screen "MTA-ALTAMC005" 1280x800, template "Plantilla-Alta-Cmp"
   Button "Botón_1" at 186,441 size 48x38; TextOff 'Incrementar'; Authorization "Operación"; PictureOff "Gráfico_3"
      on Press: SetBit("IncP5")
      on Release: ResetBit("IncP5")
   Button "Botón_2" at 186,401 size 48x38; TextOff 'Decrementar'; Authorization "Operación"; PictureOff "Gráfico_1"
      on Press: SetBit("DecP5")
      on Release: ResetBit("DecP5")
   Button "Botón_7" at 390,106 size 40x38; TextOff 'Text'; PictureOff "x"
      on Click: function_efd93a16()
   Button "Botón_8" at 310,600 size 96x35; TextOff 'Hecho'; Authorization "Administración de usuarios"
      on Press: SetTag("Varios_UltimoMantMC005_1", "HORAS5")
   TextField "Campo de texto_6" at 266,362 size 72x27; Text 'Seteada'
   TextField "Campo de texto_7" at 82,426 size 84x27; Text 'Prioridad'
   TextField "Campo de texto_8" at 362,363 size 40x27; Text 'Real'
   TextField "Campo de texto_11" at 26,343 size 158x27; Text 'Seteo de Prioridad'
   GraphicIOField "Campo ES gráfico_3" at 294,402 size 16x78; PictureList "BarraPrioridades"
      ProcessValue <- "VCMP5"
   GraphicIOField "Campo ES gráfico_5" at 374,402 size 16x78; PictureList "BarraPrioridades_1"
      ProcessValue <- "PriRealCMP5"
   SymbolicIOField "Campo ES simbólico_2" at 9,290 size 424x37; TextOff '0'; TextOn '1'; TextList "EstadoCmpAlta"
      ProcessValue <- "Est5"
      Visibility <- "MantMC005"
   TextField "Campo de texto_16" at 521,10 size 279x27; Text 'Menú Compresor ABC-5 (MC005)'
   TextField "Campo de texto_1" at 36,510 size 326x27; Text 'Tiempo de funcionamiento acumulado'
   TextField "Campo de texto_4" at 36,570 size 231x27; Text 'Próximo mantenimiento #1'
   TextField "Campo de texto_5" at 36,635 size 231x27; Text 'Próximo mantenimiento #2'
   Button "Botón_3" at 310,665 size 96x35; TextOff 'Hecho'; Authorization "Administración de usuarios"
      on Press: SetTag("Varios_UltimoMantMC005_2", "HORAS5")
   IOField "Campo ES_4" at 574,609 size 96x32; FormatPattern 99; Unit  min
      ProcessValue <- "DB-PurgaComAlta_Toff_PurgaABC5"
   IOField "Campo ES_5" at 574,654 size 96x32; FormatPattern 99; Unit  seg
      ProcessValue <- "DB-PurgaComAlta_Ton_PurgaABC5"
   TextField "Campo de texto_2" at 459,613 size 97x27; Text 'Tiempo Off'
   TextField "Campo de texto_3" at 459,655 size 96x27; Text 'Tiempo On'
   Switch "Interruptor_2" at 459,548 size 120x40; TextOff 'OFF'; CaptionText 'Switch'; TextOn 'ON'
      ProcessValue <- "DB-PurgaComAlta_Habil_PurgaABC5"
   Button "Botón_4" at 595,548 size 80x40; TextOff 'Prueba'
      on Press: SetBit("DB-PurgaComAlta_Prueba_PurgaABC5")
      on Release: ResetBit("DB-PurgaComAlta_Prueba_PurgaABC5")
      Appearance <- "MC005_EVP"
      ObjectEnable <- "MC005_EVP"
   TextField "Campo de texto_9" at 456,510 size 131x27; Text 'Ciclo de Purga:'
   GraphicIOField "Campo ES gráfico_2" at 10,280 size 422x6; PictureList "Indicador"
      ProcessValue <- "AnimMotorMC005"
   SymbolicIOField "Campo ES simbólico_4" at 19,246 size 290x21; TextOff '0'; TextOn '1'; TextList "EstadoMotor"
      ProcessValue <- "AnimMotorMC005"
   Button "Botón_6" at 13,154 size 88x62; TextOff 'ABC 5'
   Switch "Interruptor_1" at 150,167 size 37x37; TextOn '1'; TextOff '0'; CaptionText 'Switch'; PictureOff "A2"; Authorization "Operación"; PictureOn "A"
      ProcessValue <- "Auto5"
      Visibility <- "MantMC005"
   ScreenModuleView "Faceplate_6_1" at 342,236 size 76x34; ScreenModuleType ""
      Guid_{11997190-52606} <- "IndV5"
      Guid_{11997190-52610} <- "IndR5"
      Guid_{11997190-52608} <- "IndVparp5"
   ScreenModuleView "Faceplate_7_1" at 213,158 size 207x70
      Guid_{11997190-23983} <- "ParadaMC005"
      Guid_{11997190-23981} <- "MarchaMC005"
      Guid_{11997190-90329} <- "ForzarParada5"
      Guid_{11997190-180841} <- "MantMC005"
      Guid_{11997190-89807} <- "SPOFFF5"
      Guid_{11997190-89795} <- "ForzandoMarcha5"
      Guid_{11997190-90325} <- "MarchaMC005"
      Guid_{11997190-88662} <- "MarchaOK5"
      Guid_{11997190-23985} <- "AnimMenuMC005"
      Guid_{11997190-89805} <- "SPONF5"
   IOField "Campo ES_7" at 24,535 size 173x35; Authorization "Administración de usuarios"; FormatPattern 999999999; Unit  hs
      ProcessValue <- "HORAS5"
      Appearance <- "EstadoMantMC005"
   IOField "Campo ES_1" at 204,535 size 80x35; Authorization "Administración de usuarios"; FormatPattern 99; Unit  min
      ProcessValue <- "MIN5"
   IOField "Campo ES_2" at 24,595 size 173x35; FormatPattern 999999999; Unit  hs
      ProcessValue <- "ProxMantMC005_1"
      Appearance <- "LimiteMantMC005_1"
   IOField "Campo ES_3" at 24,660 size 173x35; FormatPattern 999999999; Unit  hs
      ProcessValue <- "ProxMantMC005_2"
      Appearance <- "LimiteMantMC005_2"

screen "MTA-Avisos" 1280x800, template "Plantilla"
   AlarmView "Visor de avisos_1" at 61,61 size 1174x631
   TextField "Campo de texto_16" at 613,9 size 54x27; Text 'Avisos'

screen "MTA-Avisos-Histórico" 1280x800, template "Plantilla"
   AlarmView "Visor de avisos_1" at 61,61 size 1174x631; AlarmLog "Fichero de avisos_MTA"
   TextField "Campo de texto_16" at 573,9 size 157x27; Text 'Histótico de Avisos'

screen "MTA-AyudaCFG1" 1280x800, template "Plantilla"
   TextField "Campo de texto_1" at 66,128 size 540x220; Text 'Cada compresor tiene su banda de presiones. Las 5 bandas para los 5 compresores se encuentran desfasadas una cantidad, determinada por el parámetro “Separación de presión entre bandas de presión de regulación”. Las posiciones de las bandas están determinadas por las prioridades. La banda de más arriba es la de Prioridad 1, y la de más abajo es la de prioridad 5. Los cambios en las prioridades que se le asignan a cada compresor no alteran el orden de las bandas de regulación. Las bandas siempre tienen el orden en función de las prioridades: la banda de más arriba es la de Prioridad 1, le sigue la 2, la 3 , la 4 y la de más abajo es la de prioridad 5.'
   TextField "Campo de texto_2" at 42,112 size 507x27; Text 'Posición de las bandas de regulación y parámetros a ajustar'
   TextField "Campo de texto_3" at 66,416 size 508x220; Text 'Cuando la presión medida se encuentre por deajo de la presión crítica inferior, cualquier compresor que se ponga en marcha comenzará a funcionar independientemente de si existen o no sopladoras encendidas. Una vez que la presión haya regresado a su nivel normal (es decir, que haya superado el valor de “Presión Crítica Superior”), los compresores regularán de manera normal, y se encenderán únicamente si existen sopladoras encendidas. La utilidad de este comportamiento, es que permite recuperar rápidamente la presión en casos tales como cuando por largo tiempo los compresores y sopladoras estuvieron apagados, y las pérdidas en las cañerías hicieron que la presión llegara a cero o a un valor cercano'
   TextField "Campo de texto_4" at 42,400 size 235x27; Text 'Utilidad de la presión crítica'
   TextField "Campo de texto_5" at 905,92 size 123x32; Text 'Banda de regulación Compresor Prioridad 1'
   TextField "Campo de texto_6" at 905,172 size 123x32; Text 'Banda de regulación Compresor Prioridad 2'
   TextField "Campo de texto_7" at 905,252 size 123x32; Text 'Banda de regulación Compresor Prioridad 3'
   TextField "Campo de texto_8" at 905,332 size 123x32; Text 'Banda de regulación Compresor Prioridad 4'
   TextField "Campo de texto_9" at 905,412 size 123x32; Text 'Banda de regulación Compresor Prioridad 5'
   TextField "Campo de texto_11" at 1148,498 size 88x32; Text 'Presión mínima para regulación'
   TextField "Campo de texto_12" at 708,557 size 128x18; Text 'Presión Crítica Superior'
   TextField "Campo de texto_13" at 708,611 size 122x18; Text 'Presión Crítica Inferior'
   TextField "Campo de texto_14" at 1162,199 size 85x46; Text 'Histéresis para regulación de presión'
   TextField "Campo de texto_15" at 658,199 size 140x46; Text 'Separación de presiones entre bandas de regulación de presión'
   Button "Botón_12" at 1089,638 size 160x49; TextOff 'Volver'
      on Click: ActivateScreen("MTA-CFGALTA", 0)
   TextField "Campo de texto_16" at 414,9 size 455x27; Text 'Ayuda: Configuración modo AUTO (Compresores Alta)'
   TextField "Campo de texto_10" at 905,492 size 123x32; Text 'Banda de regulación Compresor Prioridad 5'

screen "MTA-AyudaCmpAlta" 1280x800, template "Plantilla"
   Switch "Interruptor_1" at 1192,363 size 40x40; TextOn '1'; TextOff '0'; CaptionText 'Switch'; PictureOff "MECH2"; PictureOn "MECH1"
      ProcessValue <- "CERO"
   GraphicIOField "Campo ES gráfico_6" at 763,381 size 9x45; PictureList "BarraPrioridades"
      ProcessValue <- "VCMP3"
      Visibility <- "MantMC003"
   GraphicIOField "Campo ES gráfico_9" at 772,381 size 9x45; PictureList "BarraPrioridades_1"
      ProcessValue <- "PriRealCMP3"
      Visibility <- "MantMC003"
   GraphicView "Visor de gráficos_1" at 660,384 size 28x27; Picture "A2"
   TextField "Campo de texto_6" at 285,315 size 125x61; Text 'Estado del motor del Compresor'
   TextField "Campo de texto_10" at 413,297 size 113x61; Text 'Nombre del Compresor'
   TextField "Campo de texto_1" at 532,218 size 108x80; Text 'Estado lógico del Compresor (Programa)'
   GraphicView "Visor de gráficos_3" at 694,382 size 28x30; Picture "PilotLight_Round_GN_On_256c"
   GraphicView "Visor de gráficos_4" at 726,382 size 28x30; Picture "PilotLight_Round_RN_Off_256c"
   GraphicView "Visor de gráficos_5" at 126,91 size 28x30; Picture "PilotLight_Round_GN_Off_256c"
   GraphicView "Visor de gráficos_7" at 94,91 size 28x30; Picture "PilotLight_Round_RN_Off_256c"
   GraphicView "Visor de gráficos_8" at 126,131 size 28x30; Picture "PilotLight_Round_GN_Off_256c"
   GraphicView "Visor de gráficos_9" at 94,131 size 28x30; Picture "PilotLight_Round_RN_On_256c"
   GraphicView "Visor de gráficos_10" at 126,171 size 28x30; Picture "PilotLight_Round_GN_Off_256c"
   GraphicView "Visor de gráficos_11" at 94,171 size 28x30; Picture "PilotLight_Round_RN_On_256c"
   GraphicView "Visor de gráficos_12" at 126,211 size 28x30; Picture "PilotLight_Round_GN_On_256c"
   GraphicView "Visor de gráficos_13" at 94,211 size 28x30; Picture "PilotLight_Round_RN_Off_256c"
   GraphicView "Visor de gráficos_14" at 126,171 size 28x30; Picture "PilotLight_Round_GN_On_256c"
   GraphicIOField "Plantilla_Campo ES gráfico_5" at 897,433 size 65x60; PictureList "Motor2"
      ProcessValue <- "UNO"
   GraphicView "Visor de gráficos_2" at 924,363 size 260x142; Picture "ALTA1_1"
   GraphicView "Visor de gráficos_6" at 971,83 size 262x142; Picture "LOCAl"
   TextField "Campo de texto_7" at 607,463 size 54x42; Text 'Manual'
   TextField "Campo de texto_11" at 1067,286 size 199x76; Text 'El modo local transfiere el control del Compresor a su panel original'
   TextField "Campo de texto_12" at 1056,264 size 210x42; Text 'Activación de modo "LOCAL"'
   TextField "Campo de texto_13" at 695,98 size 210x42; Text 'Indicación de modo "LOCAL"'
   TextField "Campo de texto_16" at 926,529 size 134x42; Text 'Código de Colores'
   TextField "Campo de texto_18" at 529,9 size 241x27; Text 'Ayuda: Compresores de Alta'
   TextField "Campo de texto_3" at 703,239 size 90x80; Text 'Prioridad de arranque Seteada'
   TextField "Campo de texto_4" at 815,215 size 95x80; Text 'Prioridad de arranque Actual'
   TextField "Campo de texto_5" at 700,485 size 129x61; Text 'Horas de marcha acumuladas'
   TextField "Campo de texto_2" at 223,92 size 170x42; Text 'Deshabilitado / En Falla'
   TextField "Campo de texto_8" at 223,132 size 284x42; Text 'Habilitado y Parado / Sin requerimiento'
   TextField "Campo de texto_9" at 223,172 size 268x42; Text 'Parado con Requerimiento de Marcha'
   TextField "Campo de texto_14" at 223,212 size 122x42; Text 'En Vacío / Carga'
   TextField "Campo de texto_15" at 561,383 size 61x22; Text 'En carga'
   Button "Botón_3" at 95,559 size 280x70; TextOff 'Ayuda de Manejo'; PictureOff "x"
      on Click: ActivateScreen("MTA-AyudaCmpAlta_1", 0)
   GraphicIOField "Campo ES gráfico_4" at 421,438 size 374x6; PictureList "Indicador"
      ProcessValue <- "UNO"
   SymbolicIOField "Campo ES simbólico_4" at 440,410 size 178x21; TextOff '0'; TextOn '1'; TextList "EstadoMotor"
      ProcessValue <- "UNO"
   TextField "Campo de texto_19" at 434,377 size 66x32; Text 'ABC 2'
   IOField "Campo ES_6" at 662,413 size 85x19; FormatPattern 999999999; Unit  hs

screen "MTA-AyudaCmpAlta_1" 1280x800, template "Plantilla"
   TextField "Campo de texto_18" at 529,9 size 241x27; Text 'Ayuda: Compresores de Alta'
   TextField "Campo de texto_5" at 466,549 size 701x99; Text 'Para poder resetear las horas acumuladas de cada compresor se requiere clave de administrador. Si la cantidad máxima de horas es superada se generará un aviso y el indicador de horas se pondrá de color rojo. Para eliminar este aviso se deben resetear la cantidad de horas acumuladas, y se debería considerar la posibilidad de bajar la prioridad del compresor.'
   TextField "Campo de texto_1" at 286,362 size 72x27; Text 'Seteada'
   TextField "Campo de texto_2" at 102,426 size 84x27; Text 'Prioridad'
   TextField "Campo de texto_10" at 382,363 size 40x27; Text 'Real'
   TextField "Campo de texto_6" at 46,520 size 326x27; Text 'Tiempo de funcionamiento acumulado'
   TextField "Campo de texto_3" at 46,343 size 158x27; Text 'Seteo de Prioridad'
   Button "Botón_1" at 206,442 size 48x38; TextOff 'Incrementar'; Authorization "Operación"; PictureOff "Gráfico_3"
   Button "Botón_2" at 206,402 size 48x38; TextOff 'Decrementar'; Authorization "Operación"; PictureOff "Gráfico_1"
   Button "Botón_3" at 410,106 size 40x38; TextOff 'Text'; PictureOff "x"
      on Click: function_efd93a16()
   Button "Botón_4" at 320,558 size 96x70; TextOff 'Reset'; Authorization "Administración de usuarios"
   GraphicIOField "Campo ES gráfico_1" at 314,402 size 16x78; PictureList "BarraPrioridades"
      ProcessValue <- "VCMP2"
   GraphicIOField "Campo ES gráfico_2" at 394,402 size 16x78; PictureList "BarraPrioridades_1"
      ProcessValue <- "PriRealCMP2"
   TextField "Campo de texto_4" at 466,381 size 709x80; Text 'Para poder cambiar las prioridades de un compresor se requiere que todas las soplatoras estén desactivadas. No habrá ningúna modificación en la cantidad de compresores requeridos si el ajuste de prioridades se realiza en un tiempo menor al "Tiempo de apagado de sopladoras". Una vez terminado el ajuste el usuario debería activar nuevamente las sopladoras correspondientes.'
   TextField "Campo de texto_7" at 466,150 size 658x61; Text 'Modo MANUAL: El motor del compresor se acciona con los pulsadores de marcha y parada. El rango de presiones en el cual el compresor estará en carga debe ser seteado (On: entra en carga / Off: sale de carga) y es independiente para cada compresor.'
   TextField "Campo de texto_8" at 466,222 size 812x99; Text 'Modo AUTO: El motor del compresor va a requerir marcha de acuerdo con la cantidad de compresores necesarios para las sopladoras que estén activas. El rango de presiones en el cual el compresor estará en carga depende de su prioridad real. El compresor puede entrar en carga / requerir marcha de manera extraordinaria si la presión de la linea es menor que la "Presión Crítica" estando en modo AUTOMÁTICO.'
   TextField "Campo de texto_9" at 202,296 size 76x27; Text 'En Vacío'
   GraphicIOField "Campo ES gráfico_3" at 30,279 size 422x6; PictureList "Indicador"
      ProcessValue <- "UNO"
   SymbolicIOField "Campo ES simbólico_2" at 39,245 size 290x21; TextOff '0'; TextOn '1'; TextList "EstadoMotor"
      ProcessValue <- "UNO"
   Button "Botón_6" at 41,153 size 88x62; TextOff 'ABC 3'
   Switch "Interruptor_1" at 170,166 size 37x37; TextOn '1'; TextOff '0'; CaptionText 'Switch'; PictureOff "A2"; PictureOn "A"
      ProcessValue <- "Auto1"
      Visibility <- "MantMC002"
   ScreenModuleView "Faceplate_7_1" at 241,157 size 200x70
      Guid_{11997190-23985} <- "AnimMenuMC001"
   IOField "Campo ES_7" at 88,558 size 173x35; FormatPattern 999999999; Unit  hs
   IOField "Campo ES_1" at 103,590 size 173x35; FormatPattern 999999999; Unit  min
   GraphicView "Visor de gráficos_12" at 356,232 size 36x38; Picture "PilotLight_Round_GN_On_256c"
   GraphicView "Visor de gráficos_13" at 396,232 size 36x38; Picture "PilotLight_Round_RN_Off_256c"

screen "MTA-AyudaColores" 1280x800, template "Plantilla"
   GraphicView "Visor de gráficos_1" at 156,507 size 64x58; Picture "indAmarillo"
   GraphicView "Visor de gráficos_3" at 156,251 size 64x58; Picture "indCeleste"
   GraphicView "Visor de gráficos_4" at 156,315 size 64x58; Picture "indDorado"
   GraphicView "Visor de gráficos_5" at 156,187 size 64x58; Picture "indGris"
   GraphicView "Visor de gráficos_6" at 156,379 size 64x58; Picture "indRojo"
   GraphicView "Visor de gráficos_7" at 156,443 size 64x58; Picture "indVerde"
   TextField "Campo de texto_1" at 234,518 size 172x42; Text 'Sobrecarga de corriente'
   TextField "Campo de texto_2" at 130,112 size 233x32; Text 'Codificación de colores'
   TextField "Campo de texto_3" at 234,262 size 75x42; Text 'Habilitado'
   TextField "Campo de texto_4" at 234,326 size 431x42; Text 'Detenido (en algunos casos también significa modo manual)'
   TextField "Campo de texto_5" at 234,198 size 99x42; Text 'Deshabilitado'
   TextField "Campo de texto_6" at 234,390 size 56x42; Text 'En falla'
   TextField "Campo de texto_7" at 234,454 size 77x42; Text 'En Marcha'
   TextField "Campo de texto_8" at 130,598 size 666x58; Text 'Los colores indican los estados de los motores / compresores / secadores de manera rápida. La codificación de colores siempre está acompañada de un texto que contiene la misma información.'
   TextField "Campo de texto_9" at 130,646 size 1002x40; Text 'En algunos casos también aparecen los colores Verde Oscuro y Azul Oscuro que indican los estados de "Arrancando" y "Deteniéndose" respectivamente.'
   TextField "Campo de texto_16" at 542,9 size 200x27; Text 'Ayuda: Estados/Colores'

screen "MTA-AyudaMotores" 1280x800, template "Plantilla"
   TextField "Campo de texto_5" at 159,478 size 343x42; Text 'Representación de Motor con código de colores'
   TextField "Campo de texto_8" at 50,294 size 461x58; Text 'La Deshabilitación del motor provoca también la detención del mismo. La Habilitación del motor permite operar el pulsador de Marcha.'
   TextField "Campo de texto_9" at 882,291 size 279x58; Text 'Para poder marchar el motor es necesario que el mismo esté habilitado'
   GraphicView "Visor de gráficos_2" at 624,407 size 64x103; Picture "Bomba"
   GraphicIOField "Plantilla_Campo ES gráfico_4" at 660,481 size 81x68; PictureList "Motor2"
      ProcessValue <- "UNO"
   SymbolicIOField "Campo ES simbólico_3" at 572,220 size 220x29; TextOff '0'; TextOn '1'; TextList "EstadoMotor"
      ProcessValue <- "UNO"
   TextField "Campo de texto_10" at 575,161 size 52x23; Text 'MP013'
   TextField "Campo de texto_17" at 573,193 size 146x18; Text 'Chillers Envasado - Backup'
   ScreenModuleView "ControlMotor-NoAUTO_4" at 599,262 size 171x108
   TextField "Campo de texto_1" at 39,261 size 436x42; Text 'Habilitación/Deshabilitación del accionamiento desde el panel'
   TextField "Campo de texto_2" at 871,261 size 179x42; Text 'Orden de Marchar motor'
   TextField "Campo de texto_3" at 871,373 size 160x42; Text 'Orden de Parar motor'
   TextField "Campo de texto_4" at 119,205 size 376x42; Text 'Estado del motor (descripción del código de colores)'
   TextField "Campo de texto_6" at 871,165 size 251x23; Text 'Nombre simbólico en el programa'
   TextField "Campo de texto_7" at 871,197 size 135x42; Text 'Nombre del motor'
   TextField "Campo de texto_16" at 573,9 size 135x27; Text 'Ayuda: Motores'

screen "MTA-AyudaSecAlta" 1280x800, template "Plantilla"
   GraphicIOField "Campo ES gráfico_1" at 141,455 size 511x6; PictureList "Indicador"
      ProcessValue <- "UNO"
   GraphicIOField "Campo ES gráfico_2" at 141,639 size 511x6; PictureList "Indicador"
      ProcessValue <- "CERO"
   GraphicIOField "Campo ES gráfico_7" at 962,373 size 309x81; PictureList "Secador2"
      ProcessValue <- "UNO"
   GraphicView "Visor de gráficos_2" at 988,283 size 260x142; Picture "secador3_1"
   GraphicView "Visor de gráficos_6" at 971,83 size 262x142; Picture "secador3d_1"
   GraphicView "Visor de gráficos_1" at 318,376 size 35x35; Picture "A2"
   GraphicView "Visor de gráficos_3" at 318,562 size 35x35; Picture "A"
   GraphicView "Visor de gráficos_5" at 414,369 size 202x78; Picture "menu2"
   GraphicView "Visor de gráficos_7" at 413,552 size 231x79; Picture "menu3"
   TextField "Campo de texto_8" at 290,158 size 333x94; Text 'La Deshabilitación del Secador provoca también la detención del mismo. La Habilitación del Secador permite su operaración desde el panel.'
   TextField "Campo de texto_9" at 474,275 size 211x76; Text 'Para poder marchar el Secador es necesario que el mismo esté habilitado'
   TextField "Campo de texto_3" at 279,133 size 203x42; Text 'Habilitación/Deshabilitación'
   TextField "Campo de texto_4" at 463,245 size 192x42; Text 'Orden de Marchar Secador'
   TextField "Campo de texto_5" at 679,495 size 173x42; Text 'Orden de Parar Secador'
   TextField "Campo de texto_6" at 53,267 size 143x42; Text 'Estado del Secador'
   TextField "Campo de texto_7" at 303,295 size 54x42; Text 'Manual'
   TextField "Campo de texto_10" at 175,309 size 91x61; Text 'Nombre del Secador'
   TextField "Campo de texto_11" at 706,275 size 180x76; Text 'El modo local transfiere el control del Secador a su panel original'
   TextField "Campo de texto_12" at 695,245 size 210x42; Text 'Activación de modo "LOCAL"'
   TextField "Campo de texto_13" at 695,98 size 210x42; Text 'Indicación de modo "LOCAL"'
   TextField "Campo de texto_14" at 714,643 size 520x76; Text 'Cada Secador puede relacionar su estado con uno o dos compresores de alta. Mientras alguno de los compresores seleccionados esté en marcha, el secador se mantendrá en funcionamiento.'
   TextField "Campo de texto_15" at 703,613 size 255x42; Text 'Enclavamientos (Modo Automático)'
   TextField "Campo de texto_16" at 1062,513 size 134x42; Text 'Código de Colores'
   TextField "Campo de texto_17" at 310,487 size 38x42; Text 'Auto'
   TextField "Campo de texto_18" at 529,9 size 219x27; Text 'Ayuda: Secadores de Alta'
   TextField "Campo de texto_1" at 166,377 size 89x39; Text 'ABC 2'
   SymbolicIOField "Campo ES simbólico_1" at 168,413 size 242x21; TextOff '0'; TextOn '1'; TextList "EstadoMotor"
      ProcessValue <- "UNO"
   TextField "Campo de texto_2" at 166,561 size 89x39; Text 'ABC 2'
   SymbolicIOField "Campo ES simbólico_2" at 168,597 size 242x21; TextOff '0'; TextOn '1'; TextList "EstadoMotor"
      ProcessValue <- "CERO"
   Switch "Interruptor_1" at 928,331 size 40x40; TextOn '1'; TextOff '0'; CaptionText 'Switch'; PictureOff "MECH2"; PictureOn "MECH1"
      ProcessValue <- "CERO"

screen "MTA-AyudaSecBaja" 1280x800, template "Plantilla"
   GraphicIOField "Campo ES gráfico_3" at 626,509 size 510x6; PictureList "Indicador"
      ProcessValue <- "UNO"
   GraphicIOField "Campo ES gráfico_8" at 303,471 size 269x90; PictureList "BaseSullChico"
      ProcessValue <- "UNO"
   GraphicView "Visor de gráficos_1" at 336,357 size 201x179; Picture "secador_1"
   GraphicView "Visor de gráficos_3" at 344,125 size 201x179; Picture "Copia de secador"
   TextField "Campo de texto_11" at 50,363 size 180x76; Text 'El modo local transfiere el control del Secador a su panel original'
   TextField "Campo de texto_12" at 39,333 size 210x42; Text 'Activación de modo "LOCAL"'
   GraphicView "Visor de gráficos_5" at 917,426 size 202x78; Picture "menu2"
   TextField "Campo de texto_2" at 95,141 size 210x42; Text 'Indicación de modo "LOCAL"'
   TextField "Campo de texto_5" at 643,433 size 107x39; Text 'Sullair 1'
   TextField "Campo de texto_7" at 650,472 size 54x23; Text 'Marcha'
   TextField "Campo de texto_8" at 802,214 size 333x94; Text 'La Deshabilitación del Secador provoca también la detención del mismo. La Habilitación del Secador permite su operaración desde el panel.'
   TextField "Campo de texto_9" at 986,331 size 211x76; Text 'Para poder marchar el Secador es necesario que el mismo esté habilitado'
   TextField "Campo de texto_4" at 791,189 size 203x42; Text 'Habilitación/Deshabilitación'
   TextField "Campo de texto_10" at 975,301 size 192x42; Text 'Orden de Marchar Secador'
   TextField "Campo de texto_13" at 1031,559 size 173x42; Text 'Orden de Parar Secador'
   TextField "Campo de texto_14" at 564,558 size 143x42; Text 'Estado del Secador'
   TextField "Campo de texto_15" at 655,365 size 91x61; Text 'Nombre del Secador'
   TextField "Campo de texto_16" at 529,9 size 224x27; Text 'Ayuda: Secadores de Baja'
   Switch "Interruptor_8" at 275,422 size 40x40; TextOn '1'; TextOff '0'; CaptionText 'Switch'; PictureOff "MECH2"; PictureOn "MECH1"

screen "MTA-AyudaVentiladores" 1280x800, template "Plantilla"
   GraphicIOField "Campo ES gráfico_6" at 328,342 size 511x6; PictureList "Indicador"
      ProcessValue <- "CERO"
   TextField "Campo de texto_5" at 957,566 size 184x61; Text 'Representación de Motor con código de colores'
   TextField "Campo de texto_8" at 218,134 size 461x58; Text 'La Deshabilitación del motor provoca también la detención del mismo. La Habilitación del motor permite operarlo desde el panel.'
   TextField "Campo de texto_9" at 818,131 size 279x58; Text 'Para poder marchar el motor es necesario que el mismo esté habilitado'
   TextField "Campo de texto_1" at 207,101 size 436x42; Text 'Habilitación/Deshabilitación del accionamiento desde el panel'
   TextField "Campo de texto_2" at 807,101 size 179x42; Text 'Orden de Marchar motor'
   TextField "Campo de texto_4" at 197,542 size 250x61; Text 'Estado del motor (descripción del código de colores)'
   TextField "Campo de texto_7" at 107,251 size 135x42; Text 'Nombre del motor'
   GraphicView "Visor de gráficos_3" at 508,439 size 242x85; Picture "menu4_1"
   GraphicView "Visor de gráficos_4" at 508,253 size 226x85; Picture "menu2"
   GraphicView "Visor de gráficos_5" at 473,452 size 29x29; Picture "A"
   GraphicView "Visor de gráficos_6" at 473,268 size 29x29; Picture "A2"
   TextField "Campo de texto_12" at 957,478 size 156x61; Text 'Indicación ventilador en Marcha'
   TextField "Campo de texto_13" at 957,310 size 156x61; Text 'Indicación ventilador Detenido'
   TextField "Campo de texto_3" at 793,372 size 160x42; Text 'Orden de Parar motor'
   TextField "Campo de texto_6" at 413,638 size 729x61; Text 'Modo Automático Cada ventilador se pondrá en Marcha si la temperatura del agua sensada se encuentra por encima del valor de "On" y se apagará una vez que esté por debajo del valor de "Off"'
   TextField "Campo de texto_14" at 464,385 size 38x23; Text 'Auto'
   TextField "Campo de texto_15" at 448,209 size 54x23; Text 'Manual'
   TextField "Campo de texto_16" at 556,9 size 171x27; Text 'Ayuda: Ventiladores'
   TextField "Campo de texto_11" at 337,268 size 126x32; Text 'Ventilador 3'
   SymbolicIOField "Campo ES simbólico_1" at 339,304 size 170x21; TextOff '0'; TextOn '1'; TextList "EstadoMotor"
      ProcessValue <- "CERO"
   GraphicIOField "Campo ES gráfico_1" at 328,524 size 511x6; PictureList "Indicador"
      ProcessValue <- "UNO"
   TextField "Campo de texto_10" at 337,452 size 126x32; Text 'Ventilador 3'
   SymbolicIOField "Campo ES simbólico_2" at 339,488 size 170x21; TextOff '0'; TextOn '1'; TextList "EstadoMotor"
      ProcessValue <- "UNO"
   GraphicView "Visor de gráficos_18" at 757,262 size 71x70; Picture "Vent1"
   GraphicView "Visor de gráficos_1" at 757,446 size 71x70; Picture "Vent1"
   GraphicView "Visor de gráficos_2" at 757,446 size 71x70; Picture "Vent2"

screen "MTA-Booster" 1280x800, template "Plantilla"
   IOField "Campo ES_19" at 28,357 size 90x23; FormatPattern 999999999; Unit  hs
      ProcessValue <- "ProxMantBoost1"
      Appearance <- "LimiteMantBoost1"
   IOField "Campo ES_17" at 1109,356 size 90x23; FormatPattern 999999999; Unit  hs
      ProcessValue <- "ProxMantBoost2"
      Appearance <- "LimiteMantBoost2"
   GraphicView "Visor de gráficos_3" at 185,341 size 300x202; Picture "Booster-A"
   TextField "Campo de texto_16" at 0,10 size 1280x27; Text 'Boosters'
   GraphicIOField "Campo ES gráfico_1" at 238,431 size 64x70; PictureList "Motor Grande"
      ProcessValue <- "AnimaMotBooster"
   GraphicIOField "Campo ES gráfico_2" at 364,296 size 34x52; PictureList "Motor Chico"
      ProcessValue <- "AnimaMotBooster"
   GraphicIOField "Campo ES gráfico_3" at 208,410 size 221x101; PictureList "Hélice"
      ProcessValue <- "Booster_Conf_Marcha"
   SymbolicIOField "Campo ES simbólico_1" at 949,53 size 322x37; TextOff '0'; TextOn '1'; TextList "Presostato Ctrl"
      Appearance <- "Booster_Presost_Ctrl"
      ProcessValue <- "Booster_Presost_Ctrl"
   SymbolicIOField "Campo ES simbólico_2" at 949,95 size 321x37; TextOff '0'; TextOn '1'; TextList "Presostato de Alarma"
      ProcessValue <- "Booster_Presost_PA"
      Appearance <- "Booster_Presost_PA"
   GraphicView "Visor de gráficos_4" at 761,341 size 300x202; Picture "Booster-A"
   GraphicIOField "Campo ES gráfico_4" at 814,431 size 64x70; PictureList "Motor Grande"
      ProcessValue <- "AnimaMotBooster2"
   GraphicIOField "Campo ES gráfico_5" at 940,296 size 34x52; PictureList "Motor Chico"
      ProcessValue <- "AnimaMotBooster2"
   GraphicIOField "Campo ES gráfico_6" at 784,410 size 221x101; PictureList "Hélice"
      ProcessValue <- "Booster2_Conf_Marcha"
   GraphicView "Visor de gráficos_2" at 460,408 size 40x40; Picture "MECH2"
   GraphicView "Visor de gráficos_1" at 460,408 size 40x40; Picture "MECH1"
      Visibility <- "Booster_ModoManten"
   Button "Botón_6" at 460,408 size 40x40; TextOff 'Text'; PictureList "Mantenimiento"
      on Release: SetBit("Booster_PlsManten")
   IOField "Campo ES_1" at 217,338 size 90x23; Authorization "Administración de usuarios"; FormatPattern 999999999; Unit  hs.
      ProcessValue <- "HorasBoost1"
      Appearance <- "LimiteMantBoost1"
   IOField "Campo ES_2" at 790,338 size 90x23; Authorization "Administración de usuarios"; FormatPattern 999999999; Unit  hs.
      ProcessValue <- "HorasBoost2"
      Appearance <- "LimiteMantBoost2"
   Switch "Interruptor_2" at 361,96 size 72x40; TextOff 'No'; CaptionText 'Switch'; TextOn 'Si'
      ProcessValue <- "BoostPrHoras"
   TextField "Campo de texto_1" at 25,103 size 312x23; Text 'Control de Prioridades por horas de Marcha'
   Button "Botón_1" at 518,484 size 185x39; TextOff 'Invertir Prioridades'
      on Click: SetBit("BoostInvPMan")
      Visibility <- "BoostPrHoras"
   IOField "Campo ES_3" at 359,151 size 130x31; FormatPattern 99999; Unit  hs.
      ProcessValue <- "DifHorINVBoost"
      Visibility <- "BoostPrHoras"
   TextField "Campo de texto_2" at 241,152 size 93x23; Text 'Invertir cada'
      Visibility <- "BoostPrHoras"
   IOField "Campo ES_4" at 359,191 size 130x31; FormatPattern 99999; Unit  min.
      ProcessValue <- "TiempoAyudaON"
   TextField "Campo de texto_3" at 78,192 size 255x23; Text 'Tiempo para ayuda Booster auxiliar'
   IOField "Campo ES_5" at 359,231 size 130x31; FormatPattern 99999; Unit  seg.
      ProcessValue <- "TiempoAyudaOFF"
   TextField "Campo de texto_4" at 61,232 size 273x23; Text 'Tiempo para apagado Booster auxiliar'
   TextField "Campo de texto_5" at 187,550 size 250x27; Text 'Prioridad Marcha 2'
   TextField "Campo de texto_6" at 762,550 size 250x27; Text 'Prioridad Marcha 2'
   Button "Botón_7" at 849,639 size 100x27; TextOff 'Manual'
      on Release: SetBit("Booster2_PlsManual")
      Appearance <- "Booster2_ModoManual"
   Button "Botón_8" at 849,607 size 100x27; TextOff 'Automático'
      on Release: SetBit("Booster2_PlsAutoma")
      Appearance <- "Booster2_ModoAutoma"
   Button "Botón_9" at 960,607 size 96x27; TextOff 'Encender'; TextOn 'Encendido'
      on Release: SetBit("Booster2OrdMarcha")
      Appearance <- "Booster2_Conf_Marcha"
   Button "Botón_10" at 960,639 size 96x27; TextOff 'Detener'
      on Release: ResetBit("Booster2OrdMarcha")
   Switch "Interruptor_3" at 730,607 size 96x59; TextOff 'Deshabilitado'; CaptionText 'Habilitacion'; TextOn 'Habilitado'
      ProcessValue <- "Booster2_Habilitacion"
   GraphicView "Visor de gráficos_5" at 1036,408 size 40x40; Picture "MECH2"
   GraphicView "Visor de gráficos_6" at 1036,408 size 40x40; Picture "MECH1"
      Visibility <- "Booster2_ModoManten"
   Button "Botón_11" at 1036,408 size 40x40; TextOff 'Text'; PictureList "Mantenimiento"
      on Release: SetBit("Booster2_PlsManten")
   Button "Botón_2" at 275,639 size 96x27; TextOff 'Manual'
      on Release: SetBit("Booster_PlsManual")
      Appearance <- "Booster_ModoManual"
   Button "Botón_3" at 275,607 size 96x27; TextOff 'Automático'
      on Release: SetBit("Booster_PlsAutoma")
      Appearance <- "Booster_ModoAutoma"
   Button "Botón_5" at 384,607 size 96x27; TextOff 'Encender'; TextOn 'Encendido'
      on Release: SetBit("BoosterOrdMarcha")
      Appearance <- "Booster_Conf_Marcha"
   Button "Botón_4" at 384,639 size 96x27; TextOff 'Detener'
      on Release: ResetBit("BoosterOrdMarcha")
   Switch "Interruptor_1" at 153,607 size 96x59; TextOff 'Deshabilitado'; CaptionText 'Habilitacion'; TextOn 'Habilitado'
      ProcessValue <- "Booster_Habilitacion"
   IOField "Campo ES_6" at 217,362 size 90x23; Authorization "Administración de usuarios"; FormatPattern 99; Unit  min.
      ProcessValue <- "min_boost1"
   IOField "Campo ES_7" at 790,362 size 90x23; Authorization "Administración de usuarios"; FormatPattern 99; Unit  min.
      ProcessValue <- "MinBoost2"
   IOField "Campo ES_8" at 217,386 size 90x23; Authorization "Administración de usuarios"; FormatPattern 99; Unit  seg.
      ProcessValue <- "SegsBoost1"
   IOField "Campo ES_9" at 790,386 size 90x23; Authorization "Administración de usuarios"; FormatPattern 99; Unit  seg.
      ProcessValue <- "SegsBoost"
   IOField "Campo ES_10" at 854,140 size 90x23; FormatPattern 99.9; Unit  bar
      ObjectEnable <- "Ver_Config"
      ProcessValue <- "LimParBoostPrio1"
      Appearance <- "Ver_Config"
   IOField "Campo ES_11" at 854,169 size 90x23; FormatPattern 99.9; Unit  bar
      ObjectEnable <- "Ver_Config"
      ProcessValue <- "LimParBoostPrio2"
      Appearance <- "Ver_Config"
   IOField "Campo ES_12" at 854,198 size 90x23; FormatPattern 99.9; Unit  bar
      ProcessValue <- "Presión_Actual_Boosters"
   IOField "Campo ES_13" at 854,227 size 90x23; FormatPattern 99.9; Unit  bar
      ObjectEnable <- "Ver_Config"
      ProcessValue <- "LimArrBoostPrio1"
      Appearance <- "Ver_Config"
   IOField "Campo ES_14" at 854,256 size 90x23; FormatPattern 99.9; Unit  bar
      ObjectEnable <- "Ver_Config"
      ProcessValue <- "LimArrBoostPrio2"
      Appearance <- "Ver_Config"
   TextField "Campo de texto_7" at 949,140 size 321x139; Text 'Tipo de Control'
   TextField "Campo de texto_8" at 187,550 size 250x27; Text 'Prioridad Marcha 1'
      Visibility <- "PrioridadBoost1"
   TextField "Campo de texto_9" at 762,550 size 250x27; Text 'Prioridad Marcha 1'
      Visibility <- "PrioridadBoost2"
   Button "Botón_13" at 985,181 size 96x30; TextOff 'Presostato'
      on Click: ResetBit("Ctrl_Analógico")
      Appearance <- "Ctrl_Analógico"
   Button "Botón_14" at 1139,181 size 96x30; TextOff 'Bandas'
      on Click: SetBit("Ctrl_Analógico")
      Appearance <- "Ctrl_Analógico"
   Button "Botón_12" at 985,233 size 252x30; TextOff 'Configurar'
      on Click: InvertBit("Ver_Config")
      Appearance <- "Ver_Config"
   TrendView "Visor de curvas_1" at 5,53 size 584x236
      Visibility <- "Ver_Config"
      ValueAxis1End <- "CotaSupPresAna"
   TextField "Campo de texto_10" at 591,140 size 241x23; Text 'Límite Parada Booster Prioridad 1'
      Appearance <- "Ver_Config"
   TextField "Campo de texto_11" at 591,169 size 241x23; Text 'Límite Parada Booster Prioridad 2'
      Appearance <- "Ver_Config"
   TextField "Campo de texto_12" at 591,198 size 105x23; Text 'Presión Actual'
      Appearance <- "Ver_Config"
   TextField "Campo de texto_13" at 591,227 size 259x23; Text 'Límite Arranque Booster Prioridad 1'
      Appearance <- "Ver_Config"
   TextField "Campo de texto_14" at 591,256 size 259x23; Text 'Límite Arranque Booster Prioridad 2'
      Appearance <- "Ver_Config"
   IOField "Campo ES_15" at 854,111 size 90x23; Authorization "Administración de usuarios"; FormatPattern 999999999; Unit  hs
      ProcessValue <- "Varios_HorasMantBost2"
   TextField "Campo de texto_15" at 591,111 size 226x23; Text 'Horas Mantenimiento Booster 2'
      Appearance <- "Ver_Config"
   IOField "Campo ES_16" at 854,82 size 90x23; Authorization "Administración de usuarios"; FormatPattern 999999999; Unit  hs
      ProcessValue <- "Varios_HorasMantBost1"
   TextField "Campo de texto_17" at 591,82 size 226x23; Text 'Horas Mantenimiento Booster 1'
      Appearance <- "Ver_Config"
   Button "Botón_15" at 49,396 size 96x35; TextOff 'Hecho'; Authorization "Administración de usuarios"
      on Press: SetTag("Varios_UltimoMantBoost1", "HorasBoost1")
   TextField "Campo de texto_19" at 28,335 size 133x18; Text 'Próximo mantenimiento'
   Button "Botón_16" at 1130,395 size 96x35; TextOff 'Hecho'; Authorization "Administración de usuarios"
      on Press: SetTag("Varios_UltimoMantBoost2", "HorasBoost2")
   TextField "Campo de texto_18" at 1109,334 size 133x18; Text 'Próximo mantenimiento'

screen "MTA-CFGALTA" 1280x800, template "Plantilla"
   TextField "Campo de texto_4" at 1016,131 size 91x20; Text 'Límite Superior'
   TextField "Campo de texto_5" at 1016,163 size 84x20; Text 'Límite Inferior'
   IOField "Campo ES_4" at 1126,129 size 98x23; FormatPattern 999.99; Unit  bar
      ProcessValue <- "LimSUP1"
   IOField "Campo ES_5" at 1126,161 size 98x23; FormatPattern 999.99; Unit  bar
      ProcessValue <- "LimINF1"
   TextField "Campo de texto_1" at 49,157 size 275x27; Text 'Presión Máxima Para Regulación'
   TextField "Campo de texto_2" at 49,277 size 316x27; Text 'Histéresis Para Regulación de Presión'
   IOField "Campo ES_1" at 630,157 size 130x31; Authorization "Administración de usuarios"; FormatPattern 999.99; Unit  bar
      ProcessValue <- "PresMaX"
   IOField "Campo ES_2" at 629,277 size 130x31; Authorization "Administración de usuarios"; FormatPattern 999.99; Unit  bar
      ProcessValue <- "Hist"
   TextField "Campo de texto_6" at 49,405 size 526x27; Text 'Separación de Presión Entre Bandas de Presión de Regulación'
   IOField "Campo ES_3" at 629,405 size 130x31; Authorization "Administración de usuarios"; FormatPattern 999.99; Unit  bar
      ProcessValue <- "Delta"
   TextField "Campo de texto_7" at 902,142 size 94x27; Text 'Prioridad 1'
   TextField "Campo de texto_8" at 1016,203 size 91x20; Text 'Límite Superior'
   TextField "Campo de texto_9" at 1016,235 size 84x20; Text 'Límite Inferior'
   TextField "Campo de texto_10" at 902,214 size 94x27; Text 'Prioridad 2'
   IOField "Campo ES_6" at 1126,201 size 98x23; FormatPattern 999.99; Unit  bar
      ProcessValue <- "LimSUP2"
   IOField "Campo ES_7" at 1126,233 size 98x23; FormatPattern 999.99; Unit  bar
      ProcessValue <- "LimINF2"
   TextField "Campo de texto_11" at 1016,275 size 91x20; Text 'Límite Superior'
   TextField "Campo de texto_12" at 1016,307 size 84x20; Text 'Límite Inferior'
   TextField "Campo de texto_13" at 902,286 size 94x27; Text 'Prioridad 3'
   IOField "Campo ES_8" at 1126,273 size 98x23; FormatPattern 999.99; Unit  bar
      ProcessValue <- "LimSUP3"
   IOField "Campo ES_9" at 1126,305 size 98x23; FormatPattern 999.99; Unit  bar
      ProcessValue <- "LimINF3"
   TextField "Campo de texto_14" at 1016,347 size 91x20; Text 'Límite Superior'
   TextField "Campo de texto_15" at 1016,379 size 84x20; Text 'Límite Inferior'
   TextField "Campo de texto_16" at 902,358 size 94x27; Text 'Prioridad 4'
   IOField "Campo ES_10" at 1126,345 size 98x23; FormatPattern 999.99; Unit  bar
      ProcessValue <- "LimSUP4"
   IOField "Campo ES_11" at 1126,377 size 98x23; FormatPattern 999.99; Unit  bar
      ProcessValue <- "LimINF4"
   TextField "Campo de texto_17" at 1016,419 size 91x20; Text 'Límite Superior'
   TextField "Campo de texto_18" at 1016,451 size 84x20; Text 'Límite Inferior'
   TextField "Campo de texto_19" at 902,430 size 94x27; Text 'Prioridad 5'
   IOField "Campo ES_12" at 1126,417 size 98x23; FormatPattern 999.99; Unit  bar
      ProcessValue <- "LimSUP5"
   IOField "Campo ES_13" at 1126,449 size 98x23; FormatPattern 999.99; Unit  bar
      ProcessValue <- "LimINF5"
   Button "Botón_12" at 1076,638 size 160x49; TextOff 'Volver'
      on Click: function_efd93a16()
   TextField "Campo de texto_3" at 58,190 size 417x22; Text 'Durante la regulación de presión, nunca se superará este valor.'
   TextField "Campo de texto_20" at 58,310 size 566x40; Text 'Es la presión que debe caer para volver a encender un compresor, luego de que haya sido puesto en vacío.'
   TextField "Campo de texto_21" at 58,438 size 512x22; Text 'Es la separación entre las bandas de presión en la que regula cada compresor'
   TextField "Campo de texto_22" at 49,509 size 249x27; Text 'Histéresis para Presión Crítica'
   TextField "Campo de texto_23" at 58,542 size 542x40; Text 'Es el mismo concepto que la “Histéresis para Regulación de Presión”, pero aplicado a la presión crítica.'
   IOField "Campo ES_14" at 629,509 size 130x31; Authorization "Administración de usuarios"; FormatPattern 999.99; Unit  bar
      ProcessValue <- "HistCRT"
   TextField "Campo de texto_24" at 1016,563 size 91x20; Text 'Límite Superior'
   TextField "Campo de texto_25" at 1016,595 size 84x20; Text 'Límite Inferior'
   TextField "Campo de texto_26" at 902,574 size 55x27; Text 'Crítica'
   IOField "Campo ES_15" at 1126,561 size 98x23; FormatPattern 999.99; Unit  bar
      ProcessValue <- "LimSUPCRT"
   IOField "Campo ES_16" at 1126,593 size 98x23; FormatPattern 999.99; Unit  bar
      ProcessValue <- "LimINFCRT"
   Button "Botón_1" at 1184,68 size 48x46; TextOff '?'
      on Click: ActivateScreen("MTA-AyudaCFG1", 0)
   TextField "Campo de texto_27" at 349,9 size 585x27; Text 'Configuración de modo Automático para compresores de Alta presión'
   TextField "Campo de texto_28" at 902,502 size 94x27; Text 'Prioridad 6'
   TextField "Campo de texto_29" at 1015,491 size 91x20; Text 'Límite Superior'
   TextField "Campo de texto_30" at 1015,523 size 84x20; Text 'Límite Inferior'
   IOField "Campo ES_17" at 1125,489 size 98x23; FormatPattern 999.99; Unit  bar
      ProcessValue <- "LimSUP6"
   IOField "Campo ES_18" at 1125,521 size 98x23; FormatPattern 999.99; Unit  bar
      ProcessValue <- "LimINF6"

screen "MTA-CFGAvisosALTA" 1280x800, template "Plantilla"
   TextField "Campo de texto_1" at 71,96 size 326x27; Text 'Presión Aviso límite de presión Máxima'
   TextField "Campo de texto_2" at 683,96 size 276x27; Text 'Presión Aviso de presión elevada'
   IOField "Campo ES_1" at 499,96 size 130x31; Authorization "Administración de usuarios"; FormatPattern 999.99; Unit  bar
      ProcessValue <- "CFG-ALtaHH"
   IOField "Campo ES_2" at 1110,96 size 130x31; Authorization "Administración de usuarios"; FormatPattern 999.99; Unit  bar
      ProcessValue <- "CFG-ALtaH"
   TextField "Campo de texto_3" at 71,146 size 322x27; Text 'Presión Aviso límite de presión Mínima'
   IOField "Campo ES_4" at 498,146 size 130x31; Authorization "Administración de usuarios"; FormatPattern 999.99; Unit  bar
      ProcessValue <- "CFG-ALtaLL"
   TextField "Campo de texto_9" at 151,49 size 283x34; Text 'Avisos de ALTA PRESIÓN'
   TextField "Campo de texto_4" at 477,9 size 349x27; Text 'Configuración de avisos para Alta presión'
   TextField "Campo de texto_8" at 71,197 size 397x27; Text 'Período de mantenimiento #1 compresor ABC1'
   IOField "Campo ES_5" at 518,197 size 90x23; Authorization "Administración de usuarios"; FormatPattern 9999999; Unit  hs
      ProcessValue <- "Varios_HorasMantMC006_1"
   TextField "Campo de texto_7" at 683,197 size 397x27; Text 'Período de mantenimiento #2 compresor ABC1'
   IOField "Campo ES_6" at 1130,197 size 90x23; Authorization "Administración de usuarios"; FormatPattern 9999999; Unit  hs
      ProcessValue <- "Varios_HorasMantMC006_2"
   TextField "Campo de texto_10" at 71,246 size 397x27; Text 'Período de mantenimiento #1 compresor ABC2'
   IOField "Campo ES_7" at 518,246 size 90x23; Authorization "Administración de usuarios"; FormatPattern 9999999; Unit  hs
      ProcessValue <- "Varios_HorasMantMC001_1"
   TextField "Campo de texto_11" at 683,246 size 397x27; Text 'Período de mantenimiento #2 compresor ABC2'
   IOField "Campo ES_8" at 1130,246 size 90x23; Authorization "Administración de usuarios"; FormatPattern 9999999; Unit  hs
      ProcessValue <- "Varios_HorasMantMC001_2"
   TextField "Campo de texto_12" at 71,296 size 397x27; Text 'Período de mantenimiento #1 compresor ABC3'
   IOField "Campo ES_9" at 518,296 size 90x23; Authorization "Administración de usuarios"; FormatPattern 9999999; Unit  hs
      ProcessValue <- "Varios_HorasMantMC002_1"
   TextField "Campo de texto_14" at 71,443 size 412x27; Text 'Período de mantenimiento #1 compresor BELLIS'
   IOField "Campo ES_11" at 518,443 size 90x23; Authorization "Administración de usuarios"; FormatPattern 9999999; Unit  hs
      ProcessValue <- "Varios_HorasMantMC003_1"
   TextField "Campo de texto_15" at 683,443 size 412x27; Text 'Período de mantenimiento #2 compresor BELLIS'
   IOField "Campo ES_12" at 1130,443 size 90x23; Authorization "Administración de usuarios"; FormatPattern 9999999; Unit  hs
      ProcessValue <- "Varios_HorasMantMC003_2"
   TextField "Campo de texto_18" at 683,345 size 397x27; Text 'Período de mantenimiento #2 compresor ABC4'
   IOField "Campo ES_15" at 1130,345 size 90x23; Authorization "Administración de usuarios"; FormatPattern 9999999; Unit  hs
      ProcessValue <- "Varios_HorasMantMC004_2"
   TextField "Campo de texto_19" at 71,393 size 397x27; Text 'Período de mantenimiento #1 compresor ABC5'
   IOField "Campo ES_16" at 518,393 size 90x23; Authorization "Administración de usuarios"; FormatPattern 9999999; Unit  hs
      ProcessValue <- "Varios_HorasMantMC005_1"
   TextField "Campo de texto_20" at 683,296 size 397x27; Text 'Período de mantenimiento #2 compresor ABC3'
   IOField "Campo ES_17" at 1130,296 size 90x23; Authorization "Administración de usuarios"; FormatPattern 9999999; Unit  hs
      ProcessValue <- "Varios_HorasMantMC002_2"
   TextField "Campo de texto_17" at 71,345 size 397x27; Text 'Período de mantenimiento #1 compresor ABC4'
   IOField "Campo ES_14" at 518,345 size 90x23; Authorization "Administración de usuarios"; FormatPattern 9999999; Unit  hs
      ProcessValue <- "Varios_HorasMantMC004_1"
   TextField "Campo de texto_6" at 683,146 size 248x27; Text 'Presión Aviso de presión baja'
   IOField "Campo ES_3" at 1110,146 size 130x31; Authorization "Administración de usuarios"; FormatPattern 999.99; Unit  bar
      ProcessValue <- "CFG-ALtaL"
   TextField "Campo de texto_13" at 683,393 size 397x27; Text 'Período de mantenimiento #2 compresor ABC5'
   IOField "Campo ES_10" at 1130,393 size 90x23; Authorization "Administración de usuarios"; FormatPattern 9999999; Unit  hs
      ProcessValue <- "Varios_HorasMantMC005_2"
   TextField "Campo de texto_5" at 683,590 size 380x27; Text 'Enclavamiento de compresores por flujostato'
   Switch "Interruptor_1" at 1155,583 size 37x37; TextOn 'ON'; TextOff 'OFF'; CaptionText 'Switch'; PictureOff "icons8-unchecked-checkbox-50_1"; PictureOn "icons8-checked-checkbox-50_1"; Authorization "Administración de usuarios"
      ProcessValue <- "Enclavamientos_En1"
   TextField "Campo de texto_16" at 71,493 size 374x27; Text 'Período de mantenimiento #1 secador ABC1'
   IOField "Campo ES_13" at 518,493 size 90x23; Authorization "Administración de usuarios"; FormatPattern 9999999; Unit  hs
      ProcessValue <- "Varios_HorasMantMS050"
   TextField "Campo de texto_21" at 71,539 size 374x27; Text 'Período de mantenimiento #1 secador ABC3'
   IOField "Campo ES_18" at 518,539 size 90x23; Authorization "Administración de usuarios"; FormatPattern 9999999; Unit  hs
      ProcessValue <- "Varios_HorasMantMS051"
   TextField "Campo de texto_22" at 683,493 size 374x27; Text 'Período de mantenimiento #1 secador ABC2'
   IOField "Campo ES_19" at 1130,493 size 90x23; Authorization "Administración de usuarios"; FormatPattern 9999999; Unit  hs
      ProcessValue <- "Varios_HorasMantMS052"
   TextField "Campo de texto_23" at 683,539 size 390x27; Text 'Período de mantenimiento #1 secador Fargon'
   IOField "Campo ES_20" at 1130,539 size 90x23; Authorization "Administración de usuarios"; FormatPattern 9999999; Unit  hs
      ProcessValue <- "Varios_HorasMantMS053"
   TextField "Campo de texto_31" at 71,589 size 397x27; Text 'Temperatura crítica para enclavamiento compr'
   IOField "Campo ES_21" at 518,589 size 90x23; Authorization "Administración de usuarios"; FormatPattern 999; Unit  °C
      ProcessValue <- "DBParamCmpALTA-MTA_TempCritEnclav"
   TextField "Campo de texto_24" at 684,637 size 408x27; Text 'Enclavamiento de compresores por temperatura'
   Switch "Interruptor_2" at 1156,630 size 37x37; TextOn 'ON'; TextOff 'OFF'; CaptionText 'Switch'; PictureOff "icons8-unchecked-checkbox-50_1"; PictureOn "icons8-checked-checkbox-50_1"; Authorization "Administración de usuarios"
      ProcessValue <- "Enclavamientos_En2"